(* Logix 5000 project; controller FV vendor 1 type 14 code 217 rev 31.11; software revision 31.00; part 35 of 63 *)
(* tags used below, declared in another part *)
   Alarm_Reset : BOOL;
   Analog_Fault_No : DINT;
   Analog_Simulation_Enabled : BOOL;
   CWD : CHECKWORD_FLAGS;
   Default_Check_Time : DINT;
   Dummy : BOOL;
   FV_A_YSTNo : DINT;
   FV_A_YSTNo_PLCtoPC : DINT;
   FV_A_YSVNo : DINT;
   FV_A_YSVNo_PLCtoPC : DINT;
   FV_FV1_TTX01_AI : PlantItem;   // FV1_TTX01
   FV_FV1_TTX01_AI_RawInput : ALIAS FOR Remote_IO:10:I.Ch0Data;   // Real Analog Input , Do Not Use In Code
   FV_FV26_TTX01_AI : PlantItem;   // FV26_TTX01
   FV_FV26_TTX01_AI_RawInput : ALIAS FOR Remote_IO:8:I.Ch04Data;   // Real Analog Input , Do Not Use In Code
   FV_FV26_TTX02_AI : PlantItem;   // FV26_TTX02
   FV_FV26_TTX02_AI_RawInput : ALIAS FOR Remote_IO:8:I.Ch05Data;   // Real Analog Input , Do Not Use In Code
   FV_FV27_TTX01_AI : PlantItem;   // FV27_TTX01
   FV_FV27_TTX01_AI_RawInput : ALIAS FOR Remote_IO:8:I.Ch06Data;   // Real Analog Input , Do Not Use In Code
   FV_FV27_TTX02_AI : PlantItem;   // FV27_TTX02
   FV_FV27_TTX02_AI_RawInput : ALIAS FOR Remote_IO:8:I.Ch07Data;   // Real Analog Input , Do Not Use In Code
   FV_FV28_TTX01_AI : PlantItem;   // FV28_TTX01
   FV_FV28_TTX01_AI_RawInput : ALIAS FOR Remote_IO:8:I.Ch08Data;   // Real Analog Input , Do Not Use In Code
   FV_FV28_TTX02_AI : PlantItem;   // FV28_TTX02
   FV_FV28_TTX02_AI_RawInput : ALIAS FOR Remote_IO:8:I.Ch09Data;   // Real Analog Input , Do Not Use In Code
   FV_FV29_TTX01_AI : PlantItem;   // FV29_TTX01
   FV_FV29_TTX01_AI_RawInput : ALIAS FOR Remote_IO:8:I.Ch10Data;   // Real Analog Input , Do Not Use In Code
   FV_FV29_TTX02_AI : PlantItem;   // FV29_TTX02
   FV_FV29_TTX02_AI_RawInput : ALIAS FOR Remote_IO:8:I.Ch11Data;   // Real Analog Input , Do Not Use In Code
   FV_FV2_TTX01_AI : PlantItem;   // FV2_TTX01
   FV_FV2_TTX01_AI_RawInput : ALIAS FOR Remote_IO:10:I.Ch1Data;   // Real Analog Input , Do Not Use In Code
   FV_FV30_TTX01_AI : PlantItem;   // FV30_TTX01
   FV_FV30_TTX01_AI_RawInput : ALIAS FOR Remote_IO:8:I.Ch12Data;   // Real Analog Input , Do Not Use In Code
   FV_FV30_TTX02_AI : PlantItem;   // FV30_TTX02
   FV_FV30_TTX02_AI_RawInput : ALIAS FOR Remote_IO:8:I.Ch13Data;   // Real Analog Input , Do Not Use In Code
   FV_FV31_TTX01_AI : PlantItem;   // FV31_TTX01
   FV_FV31_TTX01_AI_RawInput : ALIAS FOR Remote_IO:8:I.Ch14Data;   // Real Analog Input , Do Not Use In Code
   FV_FV31_TTX02_AI : PlantItem;   // FV31_TTX02
   FV_FV31_TTX02_AI_RawInput : ALIAS FOR Remote_IO:8:I.Ch15Data;   // Real Analog Input , Do Not Use In Code
   FV_FV3_TTX01_AI : PlantItem;   // FV3_TTX01
   FV_FV3_TTX01_AI_RawInput : ALIAS FOR Remote_IO:10:I.Ch2Data;   // Real Analog Input , Do Not Use In Code
   FV_FV4_TTX01_AI : PlantItem;   // FV4_TTX01
   FV_FV4_TTX01_AI_RawInput : ALIAS FOR Remote_IO:10:I.Ch3Data;   // Real Analog Input , Do Not Use In Code
   FV_FV5_TTX01_AI : PlantItem;   // FV5_TTX01
   FV_FV5_TTX01_AI_RawInput : ALIAS FOR Remote_IO:10:I.Ch4Data;   // Real Analog Input , Do Not Use In Code
   FV_FV6_TTX01_AI : PlantItem;   // FV6_TTX01
   FV_FV6_TTX01_AI_RawInput : ALIAS FOR Remote_IO:10:I.Ch5Data;   // Real Analog Input , Do Not Use In Code
   FV_FV7_TTX01_AI : PlantItem;   // FV7_TTX01
   FV_FV7_TTX01_AI_RawInput : ALIAS FOR Remote_IO:10:I.Ch6Data;   // Real Analog Input , Do Not Use In Code
   FV_GLYCOL_AI : PlantItem;   // GLYCOL
   FV_GLYCOL_AI_RawInput : ALIAS FOR Remote_IO:8:I.Ch03Data;   // Real Analog Input , Do Not Use In Code
   FV_TTX_YS_001_AI : PlantItem;   // TTX_YS_001
   FV_TTX_YS_001_AI_RawInput : ALIAS FOR Remote_IO:8:I.Ch00Data;   // Real Analog Input , Do Not Use In Code
   FV_TTX_YS_002_AI : PlantItem;   // TTX_YS_002
   FV_TTX_YS_002_AI_RawInput : ALIAS FOR Remote_IO:8:I.Ch01Data;   // Real Analog Input , Do Not Use In Code
   One_Second_One_Scan : ALIAS FOR One_Second_1_scan;
   overrange_RIO_analog_value : REAL;
   underrange_RIO_analog_value : REAL;
(* FV_Common, continued *)

ROUTINE FV_A_YSTNo_PLCtoPC   (* ladder *)
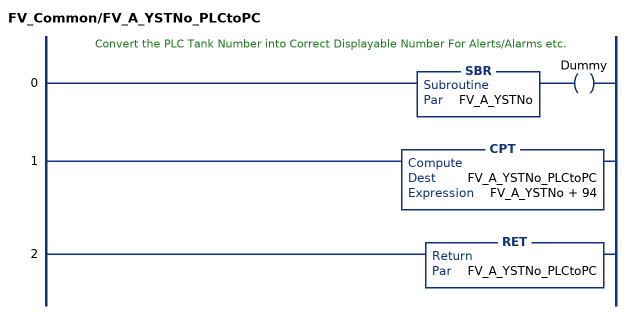
   // Convert the PLC Tank Number into Correct Displayable Number For Alerts/Alarms etc.
   0: SBR(FV_A_YSTNo)OTE(Dummy);
   1: CPT(FV_A_YSTNo_PLCtoPC,FV_A_YSTNo + 94);
   2: RET(FV_A_YSTNo_PLCtoPC);
END_ROUTINE

ROUTINE FV_A_YSVNo_PLCtoPC   (* ladder *)
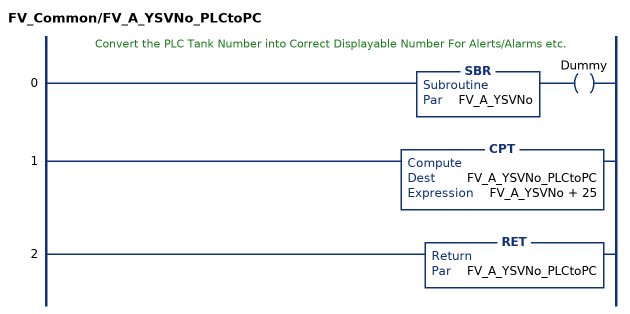
   // Convert the PLC Tank Number into Correct Displayable Number For Alerts/Alarms etc.
   0: SBR(FV_A_YSVNo)OTE(Dummy);
   1: CPT(FV_A_YSVNo_PLCtoPC,FV_A_YSVNo + 25);
   2: RET(FV_A_YSVNo_PLCtoPC);
END_ROUTINE

ROUTINE FV_Analogs   (* ladder *)
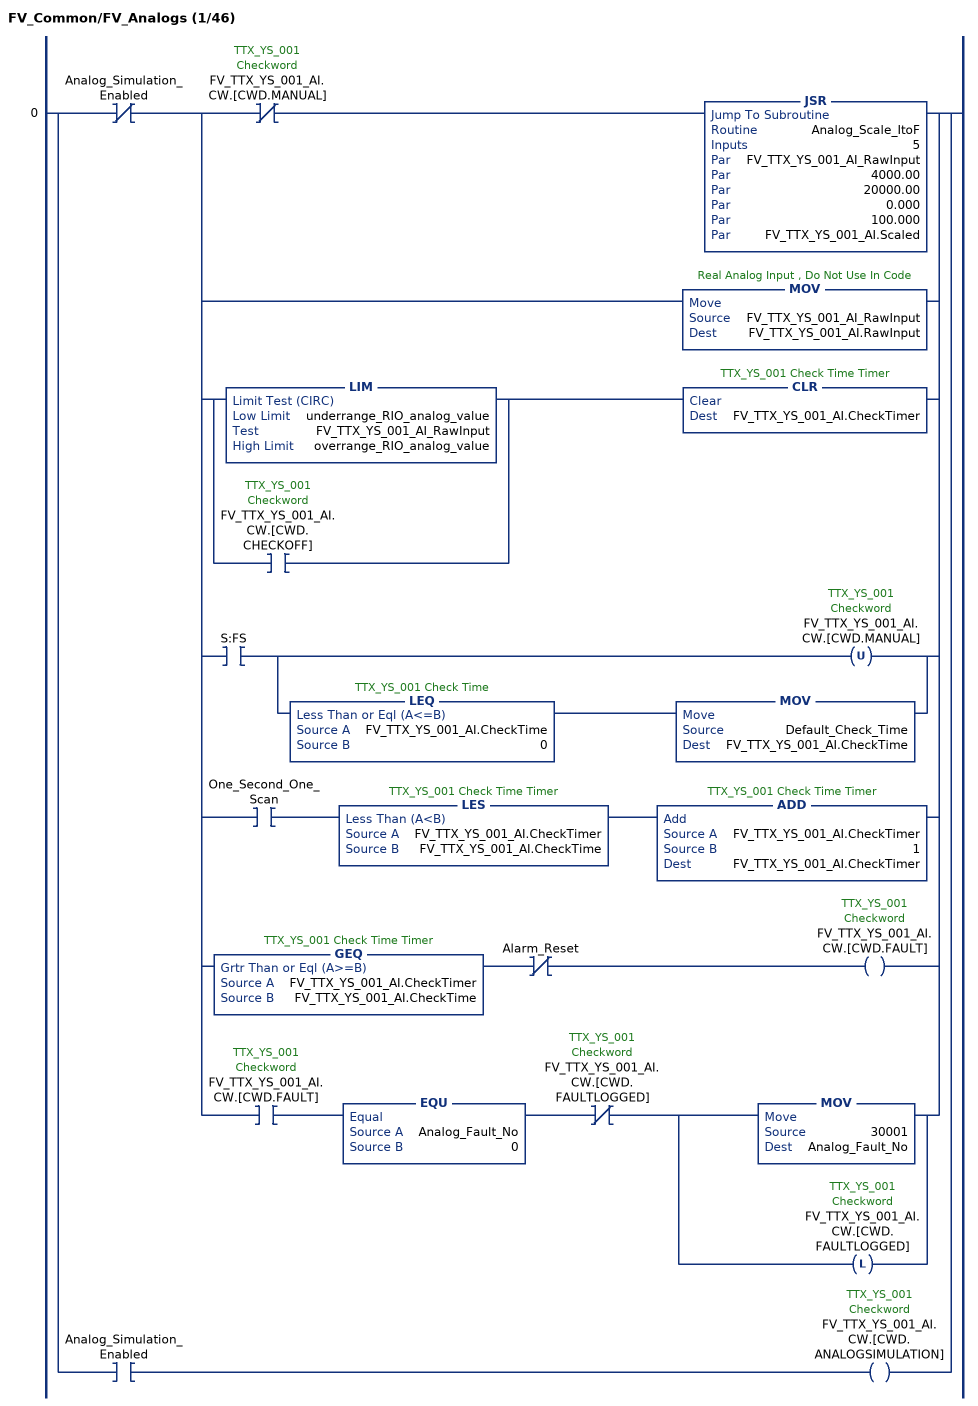
   0: [XIO(Analog_Simulation_Enabled) [XIO(FV_TTX_YS_001_AI.CW.[CWD.MANUAL]) JSR(Analog_Scale_ItoF,5,FV_TTX_YS_001_AI_RawInput,4000.00,20000.00,0.000,100.000,FV_TTX_YS_001_AI.Scaled) ,MOV(FV_TTX_YS_001_AI_RawInput,FV_TTX_YS_001_AI.RawInput) ,[LIM(underrange_RIO_analog_value,FV_TTX_YS_001_AI_RawInput,overrange_RIO_analog_value) ,XIC(FV_TTX_YS_001_AI.CW.[CWD.CHECKOFF]) ] CLR(FV_TTX_YS_001_AI.CheckTimer) ,XIC(S:FS) [OTU(FV_TTX_YS_001_AI.CW.[CWD.MANUAL]) ,LEQ(FV_TTX_YS_001_AI.CheckTime,0) MOV(Default_Check_Time,FV_TTX_YS_001_AI.CheckTime) ] ,XIC(One_Second_One_Scan) LES(FV_TTX_YS_001_AI.CheckTimer,FV_TTX_YS_001_AI.CheckTime) ADD(FV_TTX_YS_001_AI.CheckTimer,1,FV_TTX_YS_001_AI.CheckTimer) ,GEQ(FV_TTX_YS_001_AI.CheckTimer,FV_TTX_YS_001_AI.CheckTime) XIO(Alarm_Reset) OTE(FV_TTX_YS_001_AI.CW.[CWD.FAULT]) ,XIC(FV_TTX_YS_001_AI.CW.[CWD.FAULT]) EQU(Analog_Fault_No,0) XIO(FV_TTX_YS_001_AI.CW.[CWD.FAULTLOGGED]) [MOV(30001,Analog_Fault_No) ,OTL(FV_TTX_YS_001_AI.CW.[CWD.FAULTLOGGED]) ] ] ,XIC(Analog_Simulation_Enabled) OTE(FV_TTX_YS_001_AI.CW.[CWD.ANALOGSIMULATION]) ];
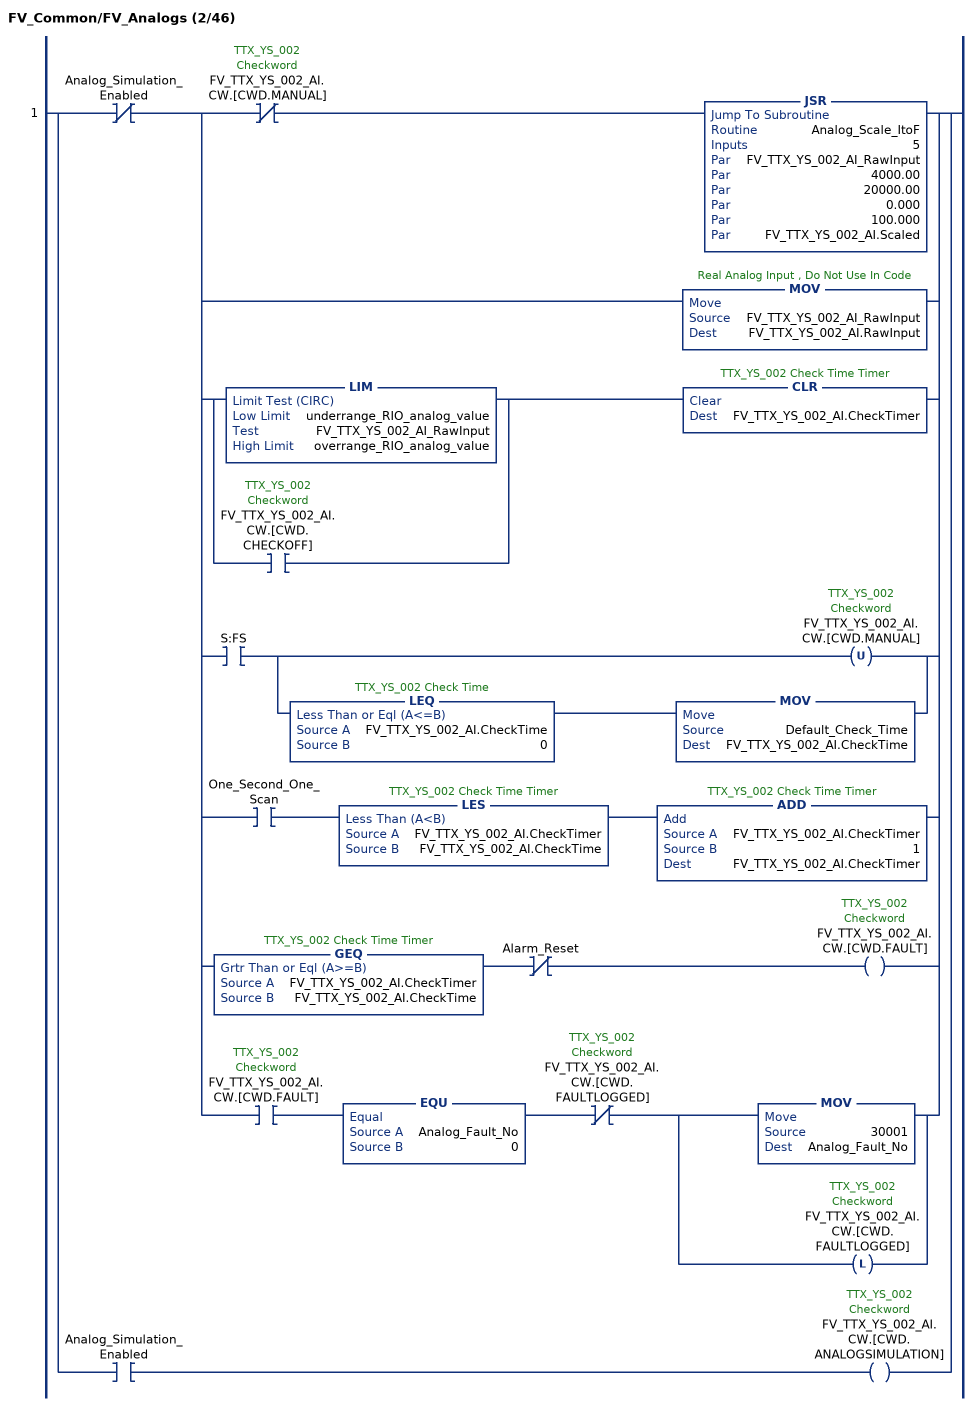
   1: [XIO(Analog_Simulation_Enabled) [XIO(FV_TTX_YS_002_AI.CW.[CWD.MANUAL]) JSR(Analog_Scale_ItoF,5,FV_TTX_YS_002_AI_RawInput,4000.00,20000.00,0.000,100.000,FV_TTX_YS_002_AI.Scaled) ,MOV(FV_TTX_YS_002_AI_RawInput,FV_TTX_YS_002_AI.RawInput) ,[LIM(underrange_RIO_analog_value,FV_TTX_YS_002_AI_RawInput,overrange_RIO_analog_value) ,XIC(FV_TTX_YS_002_AI.CW.[CWD.CHECKOFF]) ] CLR(FV_TTX_YS_002_AI.CheckTimer) ,XIC(S:FS) [OTU(FV_TTX_YS_002_AI.CW.[CWD.MANUAL]) ,LEQ(FV_TTX_YS_002_AI.CheckTime,0) MOV(Default_Check_Time,FV_TTX_YS_002_AI.CheckTime) ] ,XIC(One_Second_One_Scan) LES(FV_TTX_YS_002_AI.CheckTimer,FV_TTX_YS_002_AI.CheckTime) ADD(FV_TTX_YS_002_AI.CheckTimer,1,FV_TTX_YS_002_AI.CheckTimer) ,GEQ(FV_TTX_YS_002_AI.CheckTimer,FV_TTX_YS_002_AI.CheckTime) XIO(Alarm_Reset) OTE(FV_TTX_YS_002_AI.CW.[CWD.FAULT]) ,XIC(FV_TTX_YS_002_AI.CW.[CWD.FAULT]) EQU(Analog_Fault_No,0) XIO(FV_TTX_YS_002_AI.CW.[CWD.FAULTLOGGED]) [MOV(30001,Analog_Fault_No) ,OTL(FV_TTX_YS_002_AI.CW.[CWD.FAULTLOGGED]) ] ] ,XIC(Analog_Simulation_Enabled) OTE(FV_TTX_YS_002_AI.CW.[CWD.ANALOGSIMULATION]) ];
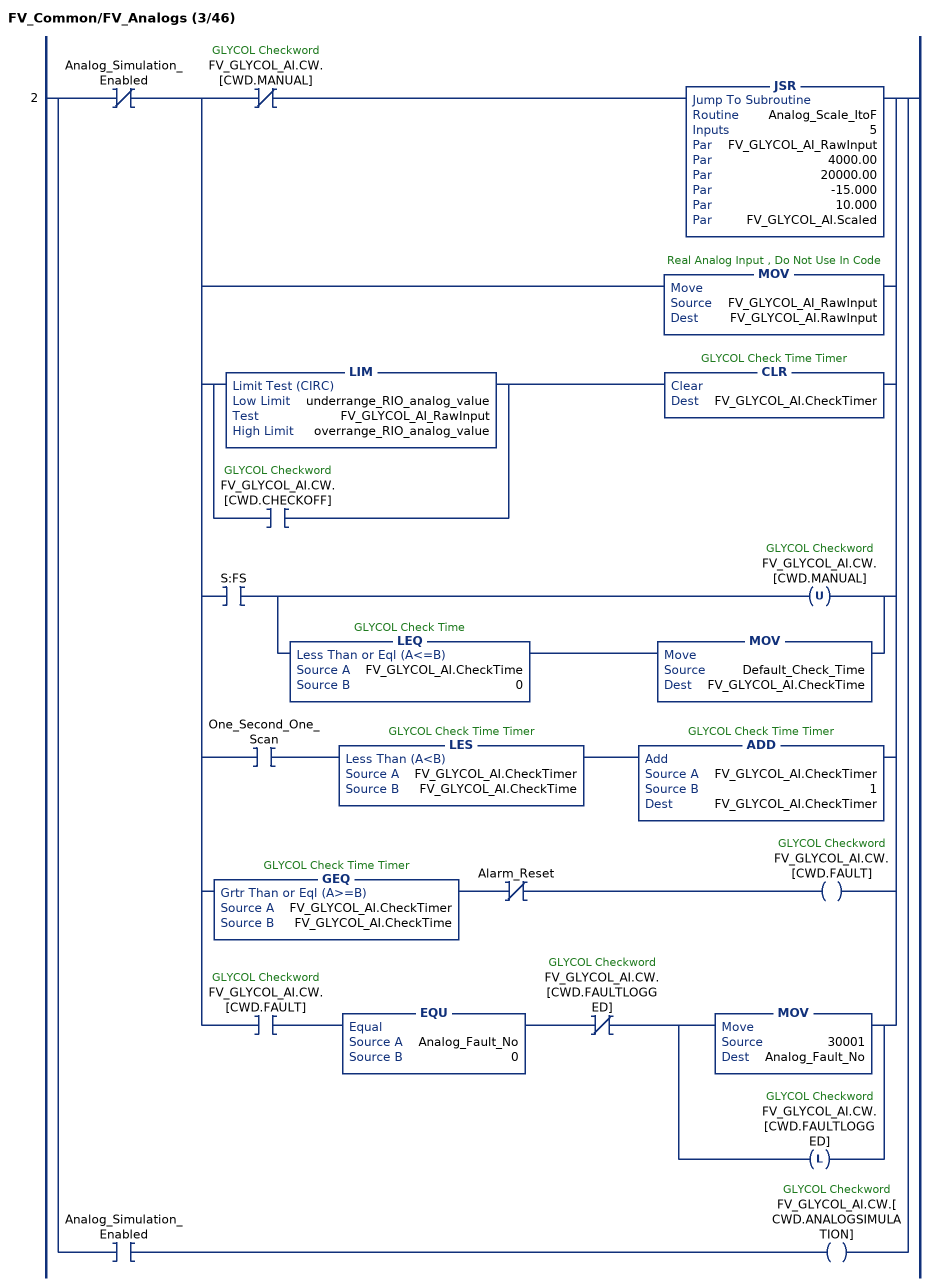
   2: [XIO(Analog_Simulation_Enabled) [XIO(FV_GLYCOL_AI.CW.[CWD.MANUAL]) JSR(Analog_Scale_ItoF,5,FV_GLYCOL_AI_RawInput,4000.00,20000.00,-15.000,10.000,FV_GLYCOL_AI.Scaled) ,MOV(FV_GLYCOL_AI_RawInput,FV_GLYCOL_AI.RawInput) ,[LIM(underrange_RIO_analog_value,FV_GLYCOL_AI_RawInput,overrange_RIO_analog_value) ,XIC(FV_GLYCOL_AI.CW.[CWD.CHECKOFF]) ] CLR(FV_GLYCOL_AI.CheckTimer) ,XIC(S:FS) [OTU(FV_GLYCOL_AI.CW.[CWD.MANUAL]) ,LEQ(FV_GLYCOL_AI.CheckTime,0) MOV(Default_Check_Time,FV_GLYCOL_AI.CheckTime) ] ,XIC(One_Second_One_Scan) LES(FV_GLYCOL_AI.CheckTimer,FV_GLYCOL_AI.CheckTime) ADD(FV_GLYCOL_AI.CheckTimer,1,FV_GLYCOL_AI.CheckTimer) ,GEQ(FV_GLYCOL_AI.CheckTimer,FV_GLYCOL_AI.CheckTime) XIO(Alarm_Reset) OTE(FV_GLYCOL_AI.CW.[CWD.FAULT]) ,XIC(FV_GLYCOL_AI.CW.[CWD.FAULT]) EQU(Analog_Fault_No,0) XIO(FV_GLYCOL_AI.CW.[CWD.FAULTLOGGED]) [MOV(30001,Analog_Fault_No) ,OTL(FV_GLYCOL_AI.CW.[CWD.FAULTLOGGED]) ] ] ,XIC(Analog_Simulation_Enabled) OTE(FV_GLYCOL_AI.CW.[CWD.ANALOGSIMULATION]) ];
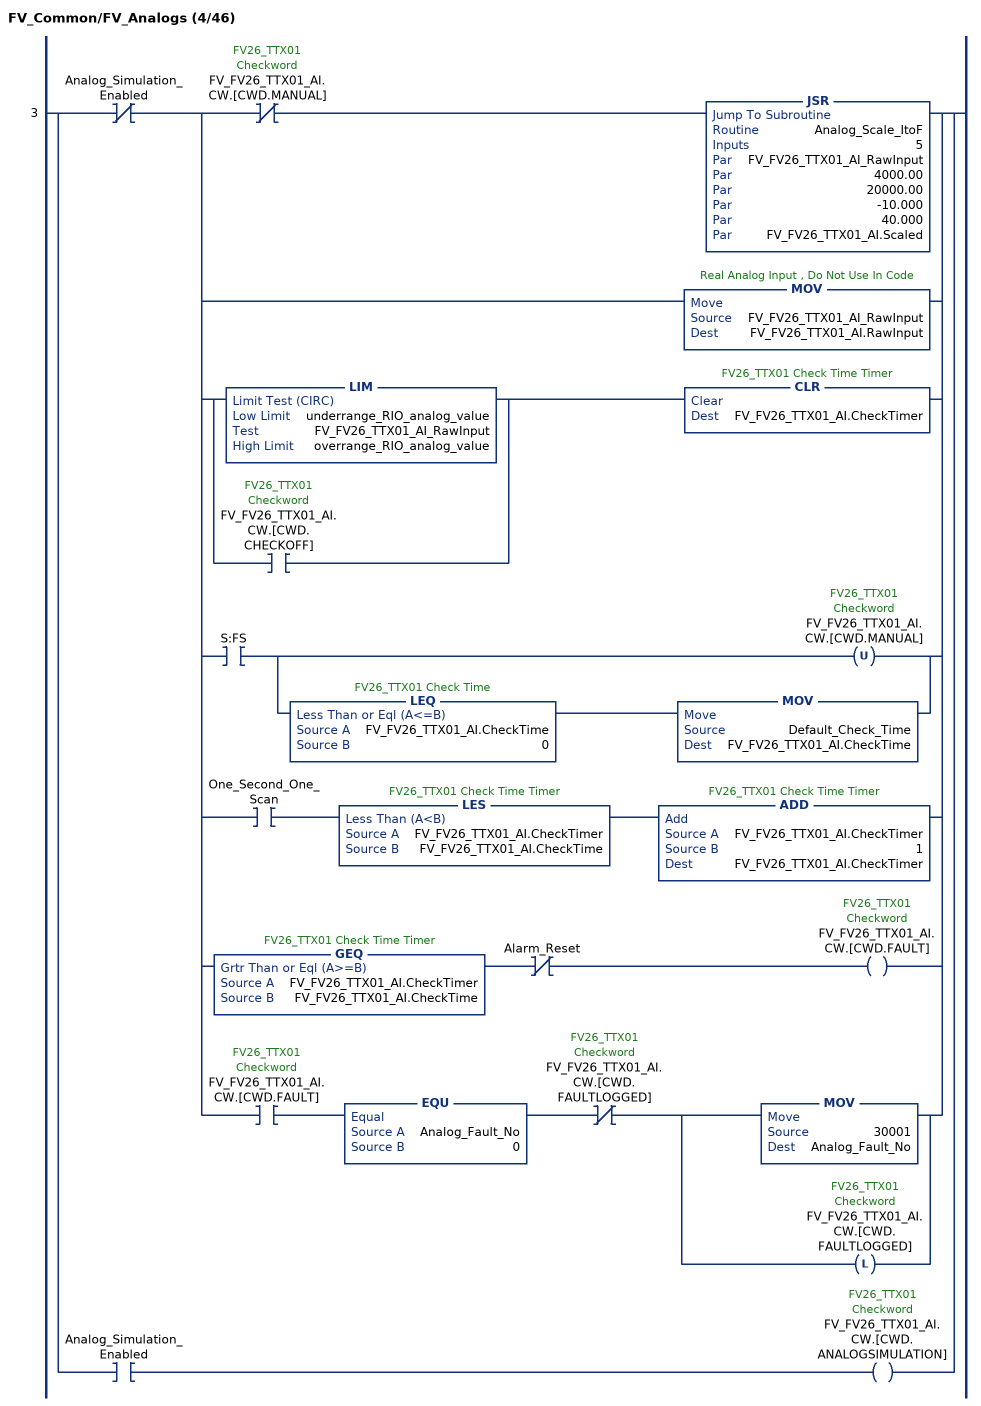
   3: [XIO(Analog_Simulation_Enabled) [XIO(FV_FV26_TTX01_AI.CW.[CWD.MANUAL]) JSR(Analog_Scale_ItoF,5,FV_FV26_TTX01_AI_RawInput,4000.00,20000.00,-10.000,40.000,FV_FV26_TTX01_AI.Scaled) ,MOV(FV_FV26_TTX01_AI_RawInput,FV_FV26_TTX01_AI.RawInput) ,[LIM(underrange_RIO_analog_value,FV_FV26_TTX01_AI_RawInput,overrange_RIO_analog_value) ,XIC(FV_FV26_TTX01_AI.CW.[CWD.CHECKOFF]) ] CLR(FV_FV26_TTX01_AI.CheckTimer) ,XIC(S:FS) [OTU(FV_FV26_TTX01_AI.CW.[CWD.MANUAL]) ,LEQ(FV_FV26_TTX01_AI.CheckTime,0) MOV(Default_Check_Time,FV_FV26_TTX01_AI.CheckTime) ] ,XIC(One_Second_One_Scan) LES(FV_FV26_TTX01_AI.CheckTimer,FV_FV26_TTX01_AI.CheckTime) ADD(FV_FV26_TTX01_AI.CheckTimer,1,FV_FV26_TTX01_AI.CheckTimer) ,GEQ(FV_FV26_TTX01_AI.CheckTimer,FV_FV26_TTX01_AI.CheckTime) XIO(Alarm_Reset) OTE(FV_FV26_TTX01_AI.CW.[CWD.FAULT]) ,XIC(FV_FV26_TTX01_AI.CW.[CWD.FAULT]) EQU(Analog_Fault_No,0) XIO(FV_FV26_TTX01_AI.CW.[CWD.FAULTLOGGED]) [MOV(30001,Analog_Fault_No) ,OTL(FV_FV26_TTX01_AI.CW.[CWD.FAULTLOGGED]) ] ] ,XIC(Analog_Simulation_Enabled) OTE(FV_FV26_TTX01_AI.CW.[CWD.ANALOGSIMULATION]) ];
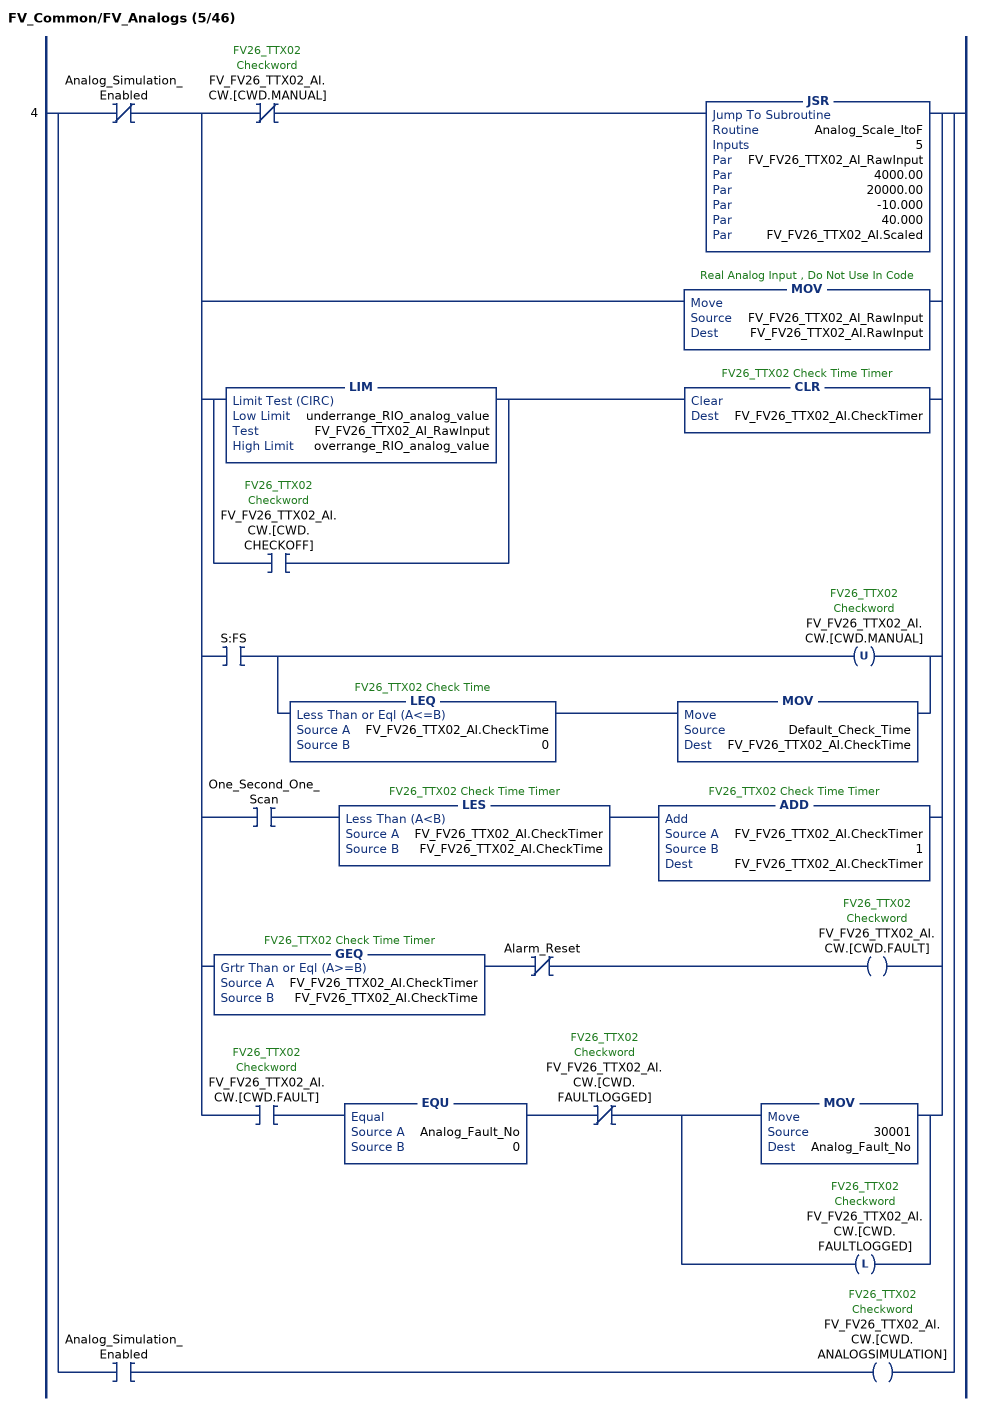
   4: [XIO(Analog_Simulation_Enabled) [XIO(FV_FV26_TTX02_AI.CW.[CWD.MANUAL]) JSR(Analog_Scale_ItoF,5,FV_FV26_TTX02_AI_RawInput,4000.00,20000.00,-10.000,40.000,FV_FV26_TTX02_AI.Scaled) ,MOV(FV_FV26_TTX02_AI_RawInput,FV_FV26_TTX02_AI.RawInput) ,[LIM(underrange_RIO_analog_value,FV_FV26_TTX02_AI_RawInput,overrange_RIO_analog_value) ,XIC(FV_FV26_TTX02_AI.CW.[CWD.CHECKOFF]) ] CLR(FV_FV26_TTX02_AI.CheckTimer) ,XIC(S:FS) [OTU(FV_FV26_TTX02_AI.CW.[CWD.MANUAL]) ,LEQ(FV_FV26_TTX02_AI.CheckTime,0) MOV(Default_Check_Time,FV_FV26_TTX02_AI.CheckTime) ] ,XIC(One_Second_One_Scan) LES(FV_FV26_TTX02_AI.CheckTimer,FV_FV26_TTX02_AI.CheckTime) ADD(FV_FV26_TTX02_AI.CheckTimer,1,FV_FV26_TTX02_AI.CheckTimer) ,GEQ(FV_FV26_TTX02_AI.CheckTimer,FV_FV26_TTX02_AI.CheckTime) XIO(Alarm_Reset) OTE(FV_FV26_TTX02_AI.CW.[CWD.FAULT]) ,XIC(FV_FV26_TTX02_AI.CW.[CWD.FAULT]) EQU(Analog_Fault_No,0) XIO(FV_FV26_TTX02_AI.CW.[CWD.FAULTLOGGED]) [MOV(30001,Analog_Fault_No) ,OTL(FV_FV26_TTX02_AI.CW.[CWD.FAULTLOGGED]) ] ] ,XIC(Analog_Simulation_Enabled) OTE(FV_FV26_TTX02_AI.CW.[CWD.ANALOGSIMULATION]) ];
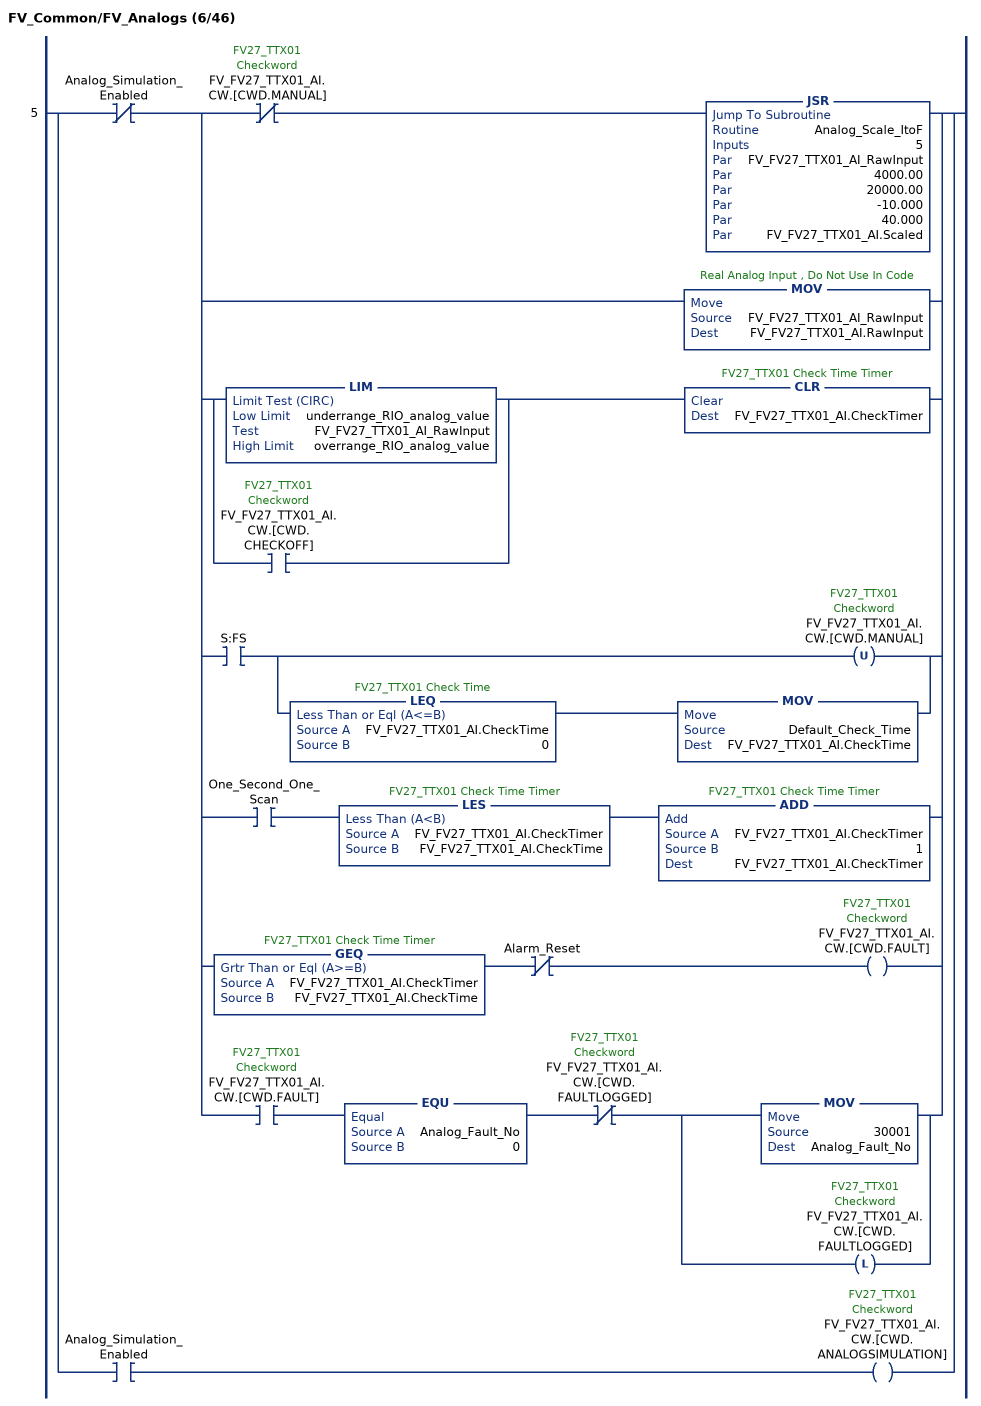
   5: [XIO(Analog_Simulation_Enabled) [XIO(FV_FV27_TTX01_AI.CW.[CWD.MANUAL]) JSR(Analog_Scale_ItoF,5,FV_FV27_TTX01_AI_RawInput,4000.00,20000.00,-10.000,40.000,FV_FV27_TTX01_AI.Scaled) ,MOV(FV_FV27_TTX01_AI_RawInput,FV_FV27_TTX01_AI.RawInput) ,[LIM(underrange_RIO_analog_value,FV_FV27_TTX01_AI_RawInput,overrange_RIO_analog_value) ,XIC(FV_FV27_TTX01_AI.CW.[CWD.CHECKOFF]) ] CLR(FV_FV27_TTX01_AI.CheckTimer) ,XIC(S:FS) [OTU(FV_FV27_TTX01_AI.CW.[CWD.MANUAL]) ,LEQ(FV_FV27_TTX01_AI.CheckTime,0) MOV(Default_Check_Time,FV_FV27_TTX01_AI.CheckTime) ] ,XIC(One_Second_One_Scan) LES(FV_FV27_TTX01_AI.CheckTimer,FV_FV27_TTX01_AI.CheckTime) ADD(FV_FV27_TTX01_AI.CheckTimer,1,FV_FV27_TTX01_AI.CheckTimer) ,GEQ(FV_FV27_TTX01_AI.CheckTimer,FV_FV27_TTX01_AI.CheckTime) XIO(Alarm_Reset) OTE(FV_FV27_TTX01_AI.CW.[CWD.FAULT]) ,XIC(FV_FV27_TTX01_AI.CW.[CWD.FAULT]) EQU(Analog_Fault_No,0) XIO(FV_FV27_TTX01_AI.CW.[CWD.FAULTLOGGED]) [MOV(30001,Analog_Fault_No) ,OTL(FV_FV27_TTX01_AI.CW.[CWD.FAULTLOGGED]) ] ] ,XIC(Analog_Simulation_Enabled) OTE(FV_FV27_TTX01_AI.CW.[CWD.ANALOGSIMULATION]) ];